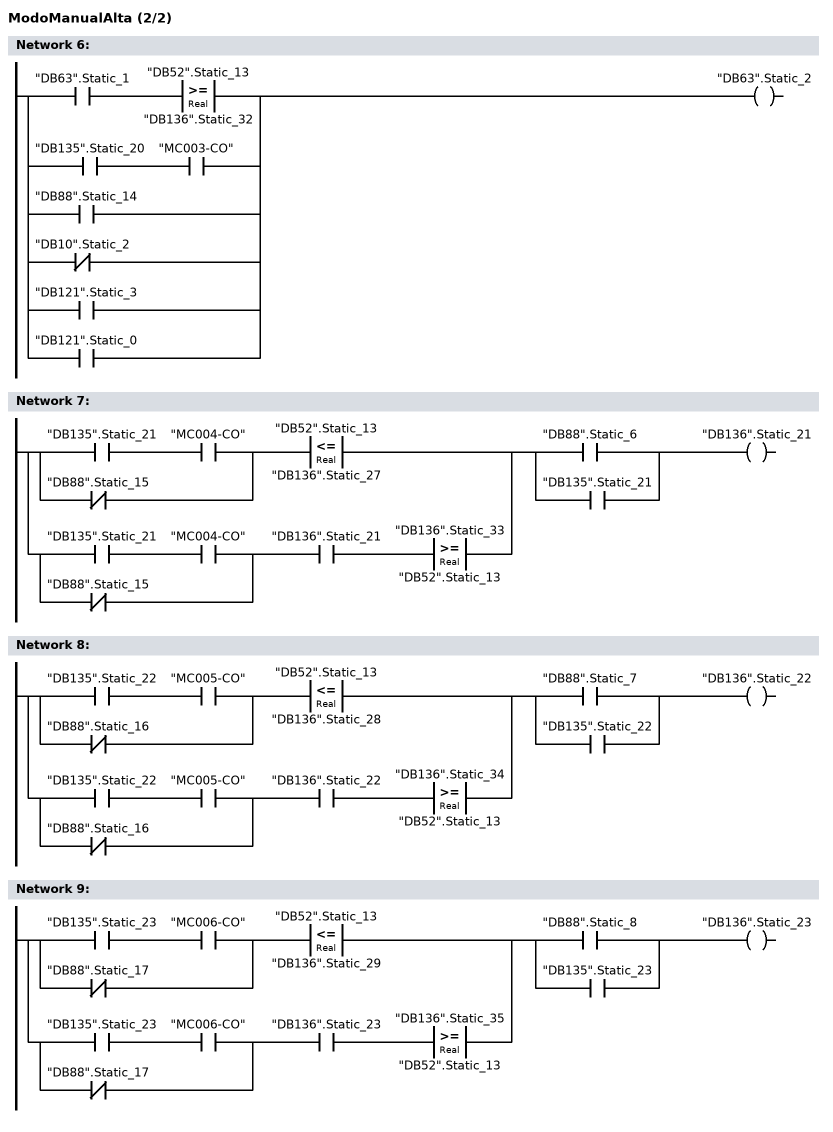
   "DB63".Static_2 := ("DB63".Static_1 AND ("DB52".Static_13 >= "DB136".Static_32)) OR "DB88".Static_14 OR ("DB135".Static_20 AND "MC003-CO") OR NOT "DB10".Static_2 OR "DB121".Static_3 OR "DB121".Static_0;
END_REGION

REGION Network 7
   "DB136".Static_21 := (((NOT "DB88".Static_15 OR ("DB135".Static_21 AND "MC004-CO")) AND ("DB52".Static_13 <= "DB136".Static_27)) OR ((NOT "DB88".Static_15 OR ("DB135".Static_21 AND "MC004-CO")) AND "DB136".Static_21 AND ("DB136".Static_33 >= "DB52".Static_13))) AND ("DB88".Static_6 OR "DB135".Static_21);
END_REGION

REGION Network 8
   "DB136".Static_22 := (((NOT "DB88".Static_16 OR ("DB135".Static_22 AND "MC005-CO")) AND ("DB52".Static_13 <= "DB136".Static_28)) OR ((NOT "DB88".Static_16 OR ("DB135".Static_22 AND "MC005-CO")) AND "DB136".Static_22 AND ("DB136".Static_34 >= "DB52".Static_13))) AND ("DB88".Static_7 OR "DB135".Static_22);
END_REGION

REGION Network 9
   "DB136".Static_23 := (((NOT "DB88".Static_17 OR ("DB135".Static_23 AND "MC006-CO")) AND ("DB52".Static_13 <= "DB136".Static_29)) OR ((NOT "DB88".Static_17 OR ("DB135".Static_23 AND "MC006-CO")) AND "DB136".Static_23 AND ("DB136".Static_35 >= "DB52".Static_13))) AND ("DB88".Static_8 OR "DB135".Static_23);
END_REGION
END_FUNCTION

// folder: Compresores/Alta/Maquina de Estados

FUNCTION "LogMaqEstGeneral" : Void   // FC35, LAD
{ S7_Optimized_Access := 'FALSE' }
VERSION : 0.1
BEGIN

REGION Network 1
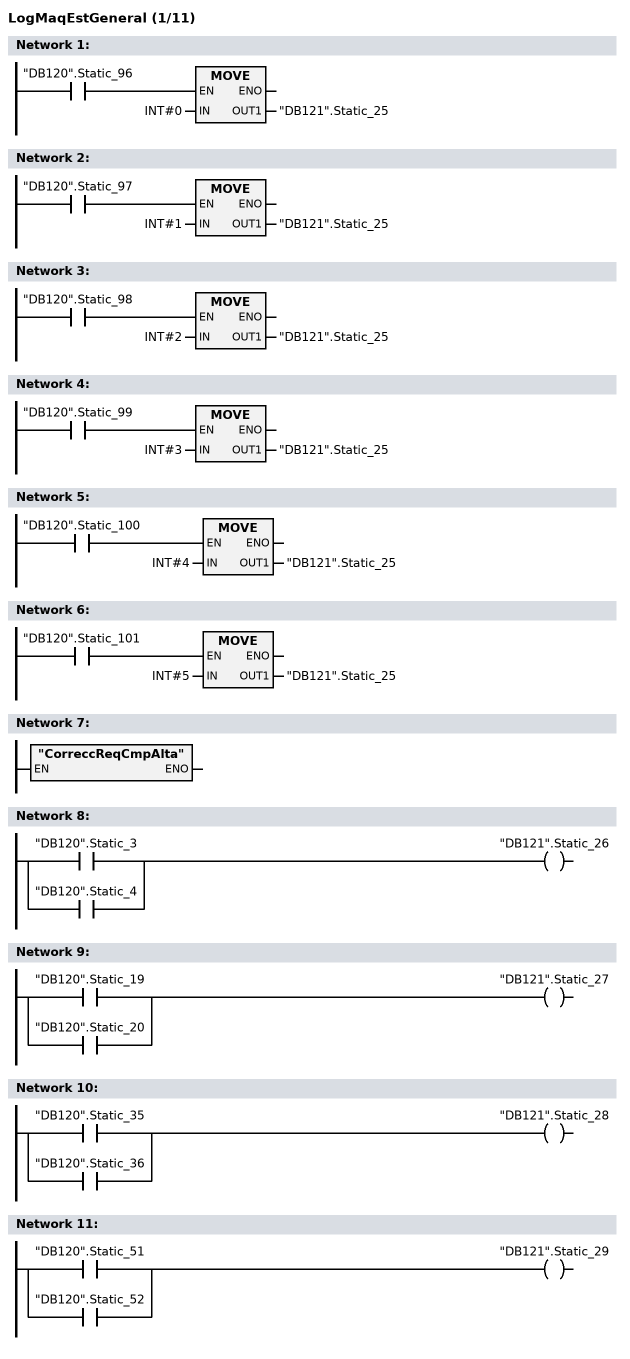
   RUNG wire#powerrail
      Contact( "DB120".Static_96 )
      { S7_GenerateENO := "TRUE" } Move(in := INT#0, out1 => "DB121".Static_25)
   END_RUNG
   // the same network as SCL:
   IF "DB120".Static_96 THEN "DB121".Static_25 := INT#0; END_IF;
END_REGION

REGION Network 2
   RUNG wire#powerrail
      Contact( "DB120".Static_97 )
      { S7_GenerateENO := "TRUE" } Move(in := INT#1, out1 => "DB121".Static_25)
   END_RUNG
   // the same network as SCL:
   IF "DB120".Static_97 THEN "DB121".Static_25 := INT#1; END_IF;
END_REGION

REGION Network 3
   RUNG wire#powerrail
      Contact( "DB120".Static_98 )
      { S7_GenerateENO := "TRUE" } Move(in := INT#2, out1 => "DB121".Static_25)
   END_RUNG
   // the same network as SCL:
   IF "DB120".Static_98 THEN "DB121".Static_25 := INT#2; END_IF;
END_REGION

REGION Network 4
   RUNG wire#powerrail
      Contact( "DB120".Static_99 )
      { S7_GenerateENO := "TRUE" } Move(in := INT#3, out1 => "DB121".Static_25)
   END_RUNG
   // the same network as SCL:
   IF "DB120".Static_99 THEN "DB121".Static_25 := INT#3; END_IF;
END_REGION

REGION Network 5
   RUNG wire#powerrail
      Contact( "DB120".Static_100 )
      { S7_GenerateENO := "TRUE" } Move(in := INT#4, out1 => "DB121".Static_25)
   END_RUNG
   // the same network as SCL:
   IF "DB120".Static_100 THEN "DB121".Static_25 := INT#4; END_IF;
END_REGION

REGION Network 6
   RUNG wire#powerrail
      Contact( "DB120".Static_101 )
      { S7_GenerateENO := "TRUE" } Move(in := INT#5, out1 => "DB121".Static_25)
   END_RUNG
   // the same network as SCL:
   IF "DB120".Static_101 THEN "DB121".Static_25 := INT#5; END_IF;
END_REGION

REGION Network 7
   RUNG wire#powerrail
      "CorreccReqCmpAlta"()
   END_RUNG
   // the same network as SCL:
   "CorreccReqCmpAlta"();
END_REGION

REGION Network 8
   RUNG wire#powerrail
      Contact( "DB120".Static_3 )
      wire#w1
      Coil( "DB121".Static_26 )
   END_RUNG
   RUNG wire#powerrail
      Contact( "DB120".Static_4 )
   END_RUNG wire#w1
   // the same network as SCL:
   "DB121".Static_26 := "DB120".Static_3 OR "DB120".Static_4;
END_REGION

REGION Network 9
   RUNG wire#powerrail
      Contact( "DB120".Static_19 )
      wire#w1
      Coil( "DB121".Static_27 )
   END_RUNG
   RUNG wire#powerrail
      Contact( "DB120".Static_20 )
   END_RUNG wire#w1
   // the same network as SCL:
   "DB121".Static_27 := "DB120".Static_19 OR "DB120".Static_20;
END_REGION

REGION Network 10
   RUNG wire#powerrail
      Contact( "DB120".Static_35 )
      wire#w1
      Coil( "DB121".Static_28 )
   END_RUNG
   RUNG wire#powerrail
      Contact( "DB120".Static_36 )
   END_RUNG wire#w1
   // the same network as SCL:
   "DB121".Static_28 := "DB120".Static_35 OR "DB120".Static_36;
END_REGION

REGION Network 11
   RUNG wire#powerrail
      Contact( "DB120".Static_51 )
      wire#w1
      Coil( "DB121".Static_29 )
   END_RUNG
   RUNG wire#powerrail
      Contact( "DB120".Static_52 )
   END_RUNG wire#w1
   // the same network as SCL:
   "DB121".Static_29 := "DB120".Static_51 OR "DB120".Static_52;
END_REGION

REGION Network 12
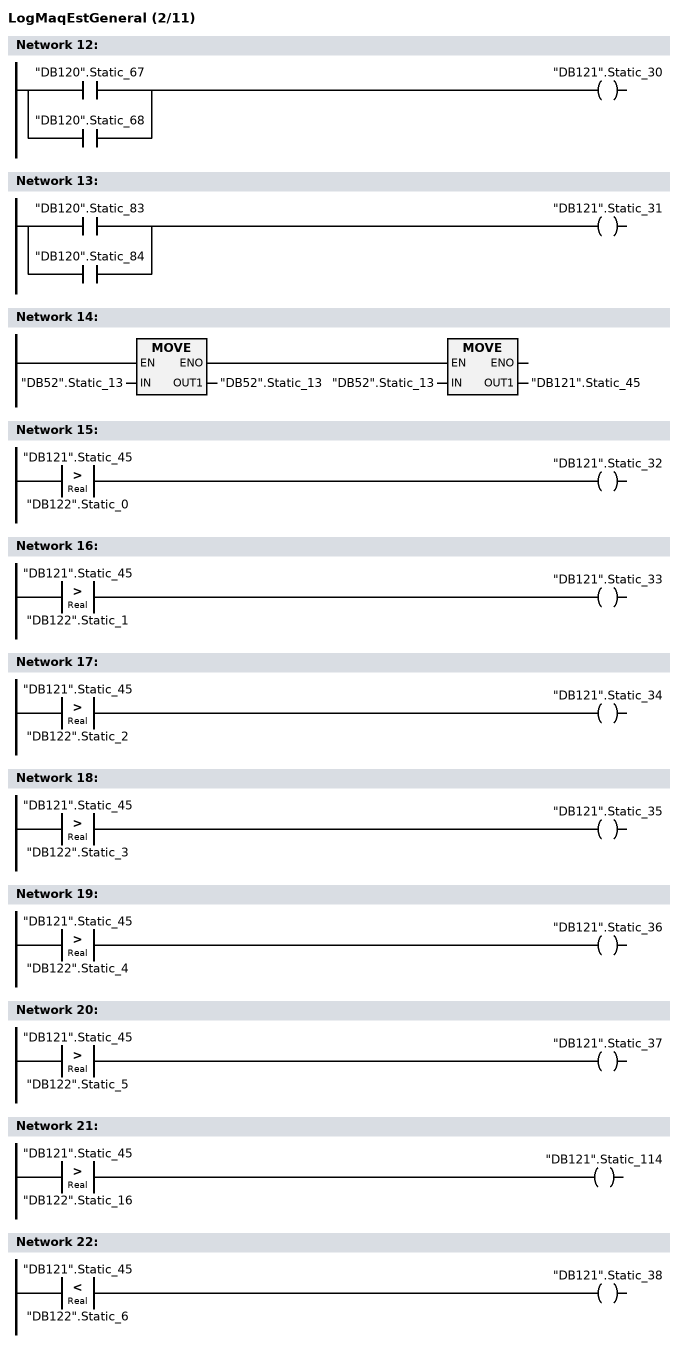
   RUNG wire#powerrail
      Contact( "DB120".Static_67 )
      wire#w1
      Coil( "DB121".Static_30 )
   END_RUNG
   RUNG wire#powerrail
      Contact( "DB120".Static_68 )
   END_RUNG wire#w1
   // the same network as SCL:
   "DB121".Static_30 := "DB120".Static_67 OR "DB120".Static_68;
END_REGION

REGION Network 13
   RUNG wire#powerrail
      Contact( "DB120".Static_83 )
      wire#w1
      Coil( "DB121".Static_31 )
   END_RUNG
   RUNG wire#powerrail
      Contact( "DB120".Static_84 )
   END_RUNG wire#w1
   // the same network as SCL:
   "DB121".Static_31 := "DB120".Static_83 OR "DB120".Static_84;
END_REGION

REGION Network 14
   RUNG wire#powerrail
      { S7_GenerateENO := "TRUE" } Move(in := "DB52".Static_13, out1 => "DB52".Static_13)
      { S7_GenerateENO := "TRUE" } Move(in := "DB52".Static_13, out1 => "DB121".Static_45)
   END_RUNG
   // the same network as SCL:
   // ENO of a box is taken as its EN; it also drops when the box reports an error
   "DB52".Static_13 := "DB52".Static_13;
   "DB121".Static_45 := "DB52".Static_13;
END_REGION

REGION Network 15
   RUNG wire#powerrail
      { S7_Templates := "SrcType := Real" } GT_Contact(in1 := "DB121".Static_45, in2 := "DB122".Static_0)
      Coil( "DB121".Static_32 )
   END_RUNG
   // the same network as SCL:
   "DB121".Static_32 := "DB121".Static_45 > "DB122".Static_0;
END_REGION

REGION Network 16
   RUNG wire#powerrail
      { S7_Templates := "SrcType := Real" } GT_Contact(in1 := "DB121".Static_45, in2 := "DB122".Static_1)
      Coil( "DB121".Static_33 )
   END_RUNG
   // the same network as SCL:
   "DB121".Static_33 := "DB121".Static_45 > "DB122".Static_1;
END_REGION

REGION Network 17
   RUNG wire#powerrail
      { S7_Templates := "SrcType := Real" } GT_Contact(in1 := "DB121".Static_45, in2 := "DB122".Static_2)
      Coil( "DB121".Static_34 )
   END_RUNG
   // the same network as SCL:
   "DB121".Static_34 := "DB121".Static_45 > "DB122".Static_2;
END_REGION

REGION Network 18
   RUNG wire#powerrail
      { S7_Templates := "SrcType := Real" } GT_Contact(in1 := "DB121".Static_45, in2 := "DB122".Static_3)
      Coil( "DB121".Static_35 )
   END_RUNG
   // the same network as SCL:
   "DB121".Static_35 := "DB121".Static_45 > "DB122".Static_3;
END_REGION

REGION Network 19
   RUNG wire#powerrail
      { S7_Templates := "SrcType := Real" } GT_Contact(in1 := "DB121".Static_45, in2 := "DB122".Static_4)
      Coil( "DB121".Static_36 )
   END_RUNG
   // the same network as SCL:
   "DB121".Static_36 := "DB121".Static_45 > "DB122".Static_4;
END_REGION

REGION Network 20
   RUNG wire#powerrail
      { S7_Templates := "SrcType := Real" } GT_Contact(in1 := "DB121".Static_45, in2 := "DB122".Static_5)
      Coil( "DB121".Static_37 )
   END_RUNG
   // the same network as SCL:
   "DB121".Static_37 := "DB121".Static_45 > "DB122".Static_5;
END_REGION

REGION Network 21
   RUNG wire#powerrail
      { S7_Templates := "SrcType := Real" } GT_Contact(in1 := "DB121".Static_45, in2 := "DB122".Static_16)
      Coil( "DB121".Static_114 )
   END_RUNG
   // the same network as SCL:
   "DB121".Static_114 := "DB121".Static_45 > "DB122".Static_16;
END_REGION

REGION Network 22
   RUNG wire#powerrail
      { S7_Templates := "SrcType := Real" } LT_Contact(in1 := "DB121".Static_45, in2 := "DB122".Static_6)
      Coil( "DB121".Static_38 )
   END_RUNG
   // the same network as SCL:
   "DB121".Static_38 := "DB121".Static_45 < "DB122".Static_6;
END_REGION

REGION Network 23
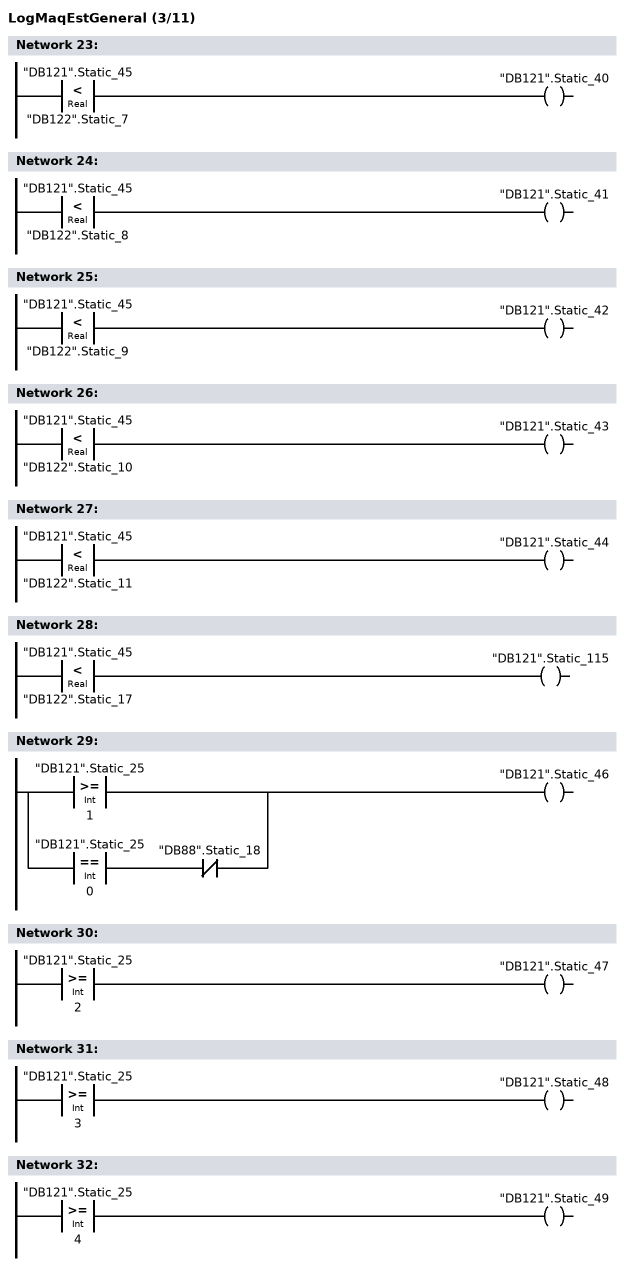
   RUNG wire#powerrail
      { S7_Templates := "SrcType := Real" } LT_Contact(in1 := "DB121".Static_45, in2 := "DB122".Static_7)
      Coil( "DB121".Static_40 )
   END_RUNG
   // the same network as SCL:
   "DB121".Static_40 := "DB121".Static_45 < "DB122".Static_7;
END_REGION

REGION Network 24
   RUNG wire#powerrail
      { S7_Templates := "SrcType := Real" } LT_Contact(in1 := "DB121".Static_45, in2 := "DB122".Static_8)
      Coil( "DB121".Static_41 )
   END_RUNG
   // the same network as SCL:
   "DB121".Static_41 := "DB121".Static_45 < "DB122".Static_8;
END_REGION

REGION Network 25
   RUNG wire#powerrail
      { S7_Templates := "SrcType := Real" } LT_Contact(in1 := "DB121".Static_45, in2 := "DB122".Static_9)
      Coil( "DB121".Static_42 )
   END_RUNG
   // the same network as SCL:
   "DB121".Static_42 := "DB121".Static_45 < "DB122".Static_9;
END_REGION

REGION Network 26
   RUNG wire#powerrail
      { S7_Templates := "SrcType := Real" } LT_Contact(in1 := "DB121".Static_45, in2 := "DB122".Static_10)
      Coil( "DB121".Static_43 )
   END_RUNG
   // the same network as SCL:
   "DB121".Static_43 := "DB121".Static_45 < "DB122".Static_10;
END_REGION

REGION Network 27
   RUNG wire#powerrail
      { S7_Templates := "SrcType := Real" } LT_Contact(in1 := "DB121".Static_45, in2 := "DB122".Static_11)
      Coil( "DB121".Static_44 )
   END_RUNG
   // the same network as SCL:
   "DB121".Static_44 := "DB121".Static_45 < "DB122".Static_11;
END_REGION

REGION Network 28
   RUNG wire#powerrail
      { S7_Templates := "SrcType := Real" } LT_Contact(in1 := "DB121".Static_45, in2 := "DB122".Static_17)
      Coil( "DB121".Static_115 )
   END_RUNG
   // the same network as SCL:
   "DB121".Static_115 := "DB121".Static_45 < "DB122".Static_17;
END_REGION

REGION Network 29
   RUNG wire#powerrail
      { S7_Templates := "SrcType := Int" } GE_Contact(in1 := "DB121".Static_25, in2 := 1)
      wire#w1
      Coil( "DB121".Static_46 )
   END_RUNG
   RUNG wire#powerrail
      { S7_Templates := "SrcType := Int" } EQ_Contact(in1 := "DB121".Static_25, in2 := 0)
      I_Contact( "DB88".Static_18 )
   END_RUNG wire#w1
   // the same network as SCL:
   "DB121".Static_46 := ("DB121".Static_25 >= 1) OR (("DB121".Static_25 = 0) AND NOT "DB88".Static_18);
END_REGION

REGION Network 30
   RUNG wire#powerrail
      { S7_Templates := "SrcType := Int" } GE_Contact(in1 := "DB121".Static_25, in2 := 2)
      Coil( "DB121".Static_47 )
   END_RUNG
   // the same network as SCL:
   "DB121".Static_47 := "DB121".Static_25 >= 2;
END_REGION

REGION Network 31
   RUNG wire#powerrail
      { S7_Templates := "SrcType := Int" } GE_Contact(in1 := "DB121".Static_25, in2 := 3)
      Coil( "DB121".Static_48 )
   END_RUNG
   // the same network as SCL:
   "DB121".Static_48 := "DB121".Static_25 >= 3;
END_REGION

REGION Network 32
   RUNG wire#powerrail
      { S7_Templates := "SrcType := Int" } GE_Contact(in1 := "DB121".Static_25, in2 := 4)
      Coil( "DB121".Static_49 )
   END_RUNG
   // the same network as SCL:
   "DB121".Static_49 := "DB121".Static_25 >= 4;
END_REGION

REGION Network 33
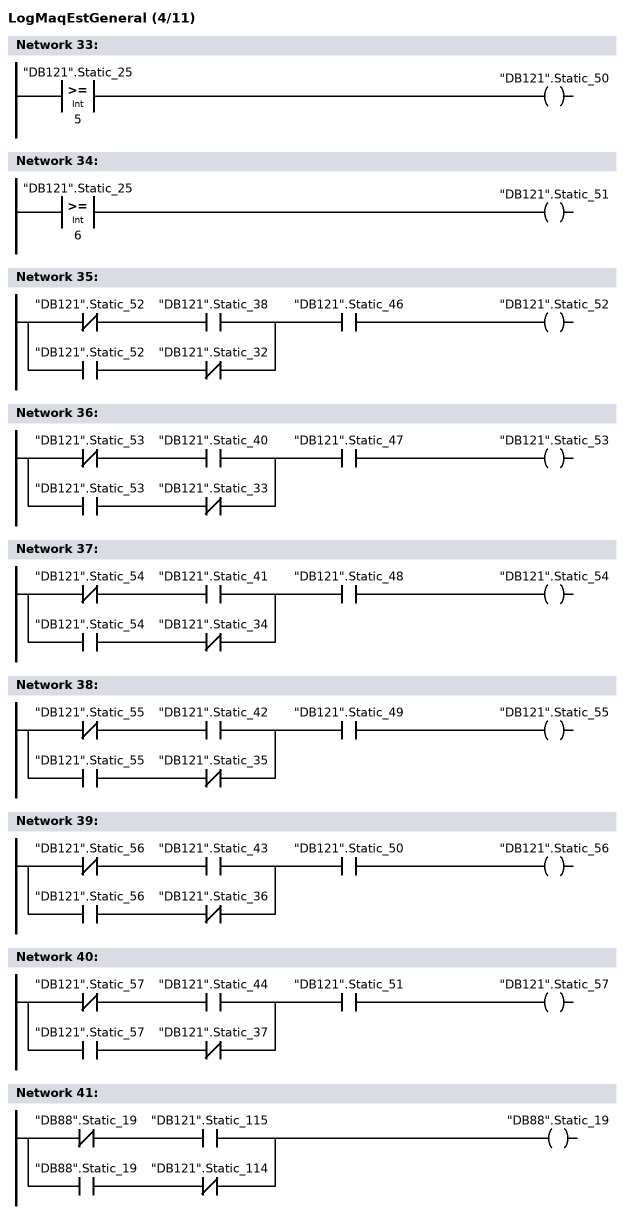
   RUNG wire#powerrail
      { S7_Templates := "SrcType := Int" } GE_Contact(in1 := "DB121".Static_25, in2 := 5)
      Coil( "DB121".Static_50 )
   END_RUNG
   // the same network as SCL:
   "DB121".Static_50 := "DB121".Static_25 >= 5;
END_REGION

REGION Network 34
   RUNG wire#powerrail
      { S7_Templates := "SrcType := Int" } GE_Contact(in1 := "DB121".Static_25, in2 := 6)
      Coil( "DB121".Static_51 )
   END_RUNG
   // the same network as SCL:
   "DB121".Static_51 := "DB121".Static_25 >= 6;
END_REGION

REGION Network 35
   RUNG wire#powerrail
      I_Contact( "DB121".Static_52 )
      Contact( "DB121".Static_38 )
      wire#w1
      Contact( "DB121".Static_46 )
      Coil( "DB121".Static_52 )
   END_RUNG
   RUNG wire#powerrail
      Contact( "DB121".Static_52 )
      I_Contact( "DB121".Static_32 )
   END_RUNG wire#w1
   // the same network as SCL:
   "DB121".Static_52 := ((NOT "DB121".Static_52 AND "DB121".Static_38) OR ("DB121".Static_52 AND NOT "DB121".Static_32)) AND "DB121".Static_46;
END_REGION

REGION Network 36
   RUNG wire#powerrail
      I_Contact( "DB121".Static_53 )
      Contact( "DB121".Static_40 )
      wire#w1
      Contact( "DB121".Static_47 )
      Coil( "DB121".Static_53 )
   END_RUNG
   RUNG wire#powerrail
      Contact( "DB121".Static_53 )
      I_Contact( "DB121".Static_33 )
   END_RUNG wire#w1
   // the same network as SCL:
   "DB121".Static_53 := ((NOT "DB121".Static_53 AND "DB121".Static_40) OR ("DB121".Static_53 AND NOT "DB121".Static_33)) AND "DB121".Static_47;
END_REGION

REGION Network 37
   RUNG wire#powerrail
      I_Contact( "DB121".Static_54 )
      Contact( "DB121".Static_41 )
      wire#w1
      Contact( "DB121".Static_48 )
      Coil( "DB121".Static_54 )
   END_RUNG
   RUNG wire#powerrail
      Contact( "DB121".Static_54 )
      I_Contact( "DB121".Static_34 )
   END_RUNG wire#w1
   // the same network as SCL:
   "DB121".Static_54 := ((NOT "DB121".Static_54 AND "DB121".Static_41) OR ("DB121".Static_54 AND NOT "DB121".Static_34)) AND "DB121".Static_48;
END_REGION

REGION Network 38
   RUNG wire#powerrail
      I_Contact( "DB121".Static_55 )
      Contact( "DB121".Static_42 )
      wire#w1
      Contact( "DB121".Static_49 )
      Coil( "DB121".Static_55 )
   END_RUNG
   RUNG wire#powerrail
      Contact( "DB121".Static_55 )
      I_Contact( "DB121".Static_35 )
   END_RUNG wire#w1
   // the same network as SCL:
   "DB121".Static_55 := ((NOT "DB121".Static_55 AND "DB121".Static_42) OR ("DB121".Static_55 AND NOT "DB121".Static_35)) AND "DB121".Static_49;
END_REGION

REGION Network 39
   RUNG wire#powerrail
      I_Contact( "DB121".Static_56 )
      Contact( "DB121".Static_43 )
      wire#w1
      Contact( "DB121".Static_50 )
      Coil( "DB121".Static_56 )
   END_RUNG
   RUNG wire#powerrail
      Contact( "DB121".Static_56 )
      I_Contact( "DB121".Static_36 )
   END_RUNG wire#w1
   // the same network as SCL:
   "DB121".Static_56 := ((NOT "DB121".Static_56 AND "DB121".Static_43) OR ("DB121".Static_56 AND NOT "DB121".Static_36)) AND "DB121".Static_50;
END_REGION

REGION Network 40
   RUNG wire#powerrail
      I_Contact( "DB121".Static_57 )
      Contact( "DB121".Static_44 )
      wire#w1
      Contact( "DB121".Static_51 )
      Coil( "DB121".Static_57 )
   END_RUNG
   RUNG wire#powerrail
      Contact( "DB121".Static_57 )
      I_Contact( "DB121".Static_37 )
   END_RUNG wire#w1
   // the same network as SCL:
   "DB121".Static_57 := ((NOT "DB121".Static_57 AND "DB121".Static_44) OR ("DB121".Static_57 AND NOT "DB121".Static_37)) AND "DB121".Static_51;
END_REGION

REGION Network 41
   RUNG wire#powerrail
      I_Contact( "DB88".Static_19 )
      Contact( "DB121".Static_115 )
      wire#w1
      Coil( "DB88".Static_19 )
   END_RUNG
   RUNG wire#powerrail
      Contact( "DB88".Static_19 )
      I_Contact( "DB121".Static_114 )
   END_RUNG wire#w1
   // the same network as SCL:
   "DB88".Static_19 := (NOT "DB88".Static_19 AND "DB121".Static_115) OR ("DB88".Static_19 AND NOT "DB121".Static_114);
END_REGION

REGION Network 42
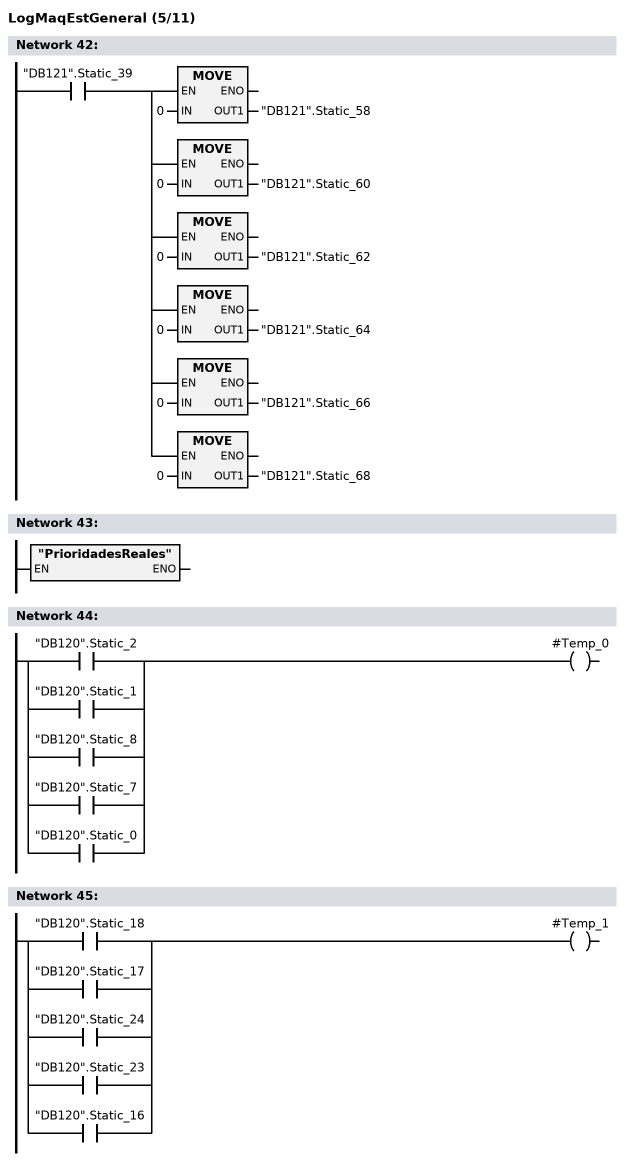
   RUNG wire#powerrail
      Contact( "DB121".Static_39 )
      wire#w1
      { S7_GenerateENO := "TRUE" } Move(in := 0, out1 => "DB121".Static_58)
   END_RUNG
   RUNG wire#w1
      { S7_GenerateENO := "TRUE" } Move(in := 0, out1 => "DB121".Static_60)
   END_RUNG
   RUNG wire#w1
      { S7_GenerateENO := "TRUE" } Move(in := 0, out1 => "DB121".Static_62)
   END_RUNG
   RUNG wire#w1
      { S7_GenerateENO := "TRUE" } Move(in := 0, out1 => "DB121".Static_64)
   END_RUNG
   RUNG wire#w1
      { S7_GenerateENO := "TRUE" } Move(in := 0, out1 => "DB121".Static_66)
   END_RUNG
   RUNG wire#w1
      { S7_GenerateENO := "TRUE" } Move(in := 0, out1 => "DB121".Static_68)
   END_RUNG
   // the same network as SCL:
   IF "DB121".Static_39 THEN
       "DB121".Static_58 := 0;
       "DB121".Static_60 := 0;
       "DB121".Static_62 := 0;
       "DB121".Static_64 := 0;
       "DB121".Static_66 := 0;
       "DB121".Static_68 := 0;
   END_IF;
END_REGION

REGION Network 43
   RUNG wire#powerrail
      "PrioridadesReales"()
   END_RUNG
   // the same network as SCL:
   "PrioridadesReales"();
END_REGION

REGION Network 44
   RUNG wire#powerrail
      Contact( "DB120".Static_2 )
      wire#w1
      Coil( #Temp_0 )
   END_RUNG
   RUNG wire#powerrail
      Contact( "DB120".Static_1 )
   END_RUNG wire#w1
   RUNG wire#powerrail
      Contact( "DB120".Static_8 )
   END_RUNG wire#w1
   RUNG wire#powerrail
      Contact( "DB120".Static_7 )
   END_RUNG wire#w1
   RUNG wire#powerrail
      Contact( "DB120".Static_0 )
   END_RUNG wire#w1
   // the same network as SCL:
   #Temp_0 := "DB120".Static_2 OR "DB120".Static_1 OR "DB120".Static_8 OR "DB120".Static_7 OR "DB120".Static_0;
END_REGION

REGION Network 45
   RUNG wire#powerrail
      Contact( "DB120".Static_18 )
      wire#w1
      Coil( #Temp_1 )
   END_RUNG
   RUNG wire#powerrail
      Contact( "DB120".Static_17 )
   END_RUNG wire#w1
   RUNG wire#powerrail
      Contact( "DB120".Static_24 )
   END_RUNG wire#w1
   RUNG wire#powerrail
      Contact( "DB120".Static_23 )
   END_RUNG wire#w1
   RUNG wire#powerrail
      Contact( "DB120".Static_16 )
   END_RUNG wire#w1
   // the same network as SCL:
   #Temp_1 := "DB120".Static_18 OR "DB120".Static_17 OR "DB120".Static_24 OR "DB120".Static_23 OR "DB120".Static_16;
END_REGION

REGION Network 46
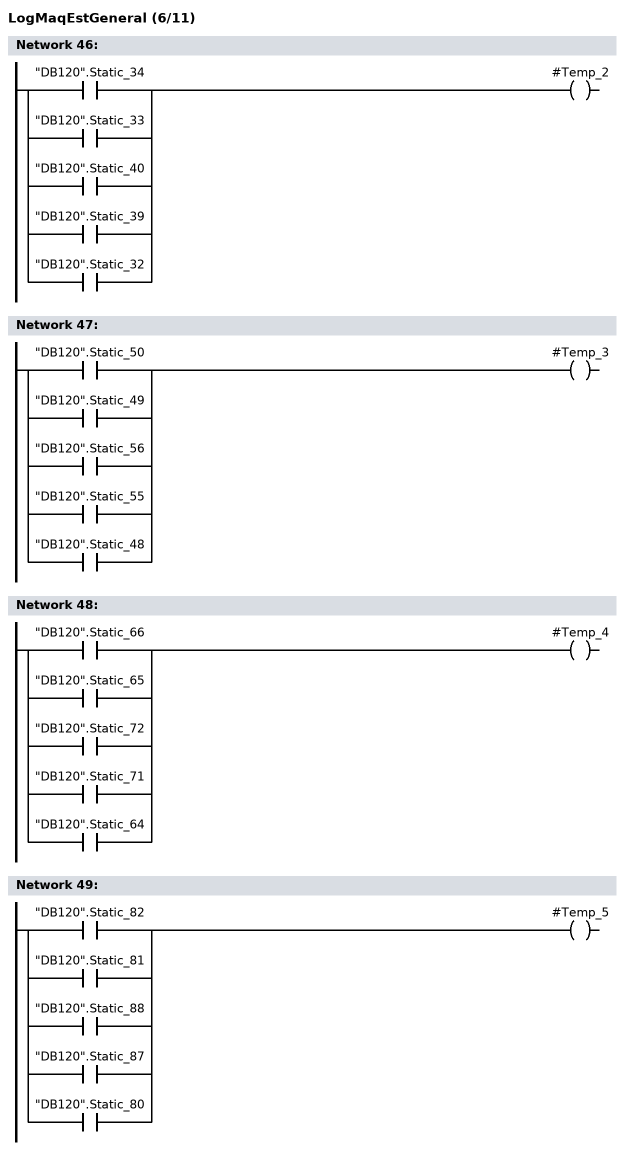
   RUNG wire#powerrail
      Contact( "DB120".Static_34 )
      wire#w1
      Coil( #Temp_2 )
   END_RUNG
   RUNG wire#powerrail
      Contact( "DB120".Static_33 )
   END_RUNG wire#w1
   RUNG wire#powerrail
      Contact( "DB120".Static_40 )
   END_RUNG wire#w1
   RUNG wire#powerrail
      Contact( "DB120".Static_39 )
   END_RUNG wire#w1
   RUNG wire#powerrail
      Contact( "DB120".Static_32 )
   END_RUNG wire#w1
   // the same network as SCL:
   #Temp_2 := "DB120".Static_34 OR "DB120".Static_33 OR "DB120".Static_40 OR "DB120".Static_39 OR "DB120".Static_32;
END_REGION

REGION Network 47
   RUNG wire#powerrail
      Contact( "DB120".Static_50 )
      wire#w1
      Coil( #Temp_3 )
   END_RUNG
   RUNG wire#powerrail
      Contact( "DB120".Static_49 )
   END_RUNG wire#w1
   RUNG wire#powerrail
      Contact( "DB120".Static_56 )
   END_RUNG wire#w1
   RUNG wire#powerrail
      Contact( "DB120".Static_55 )
   END_RUNG wire#w1
   RUNG wire#powerrail
      Contact( "DB120".Static_48 )
   END_RUNG wire#w1
   // the same network as SCL:
   #Temp_3 := "DB120".Static_50 OR "DB120".Static_49 OR "DB120".Static_56 OR "DB120".Static_55 OR "DB120".Static_48;
END_REGION

REGION Network 48
   RUNG wire#powerrail
      Contact( "DB120".Static_66 )
      wire#w1
      Coil( #Temp_4 )
   END_RUNG
   RUNG wire#powerrail
      Contact( "DB120".Static_65 )
   END_RUNG wire#w1
   RUNG wire#powerrail
      Contact( "DB120".Static_72 )
   END_RUNG wire#w1
   RUNG wire#powerrail
      Contact( "DB120".Static_71 )
   END_RUNG wire#w1
   RUNG wire#powerrail
      Contact( "DB120".Static_64 )
   END_RUNG wire#w1
   // the same network as SCL:
   #Temp_4 := "DB120".Static_66 OR "DB120".Static_65 OR "DB120".Static_72 OR "DB120".Static_71 OR "DB120".Static_64;
END_REGION

REGION Network 49
   RUNG wire#powerrail
      Contact( "DB120".Static_82 )
      wire#w1
      Coil( #Temp_5 )
   END_RUNG
   RUNG wire#powerrail
      Contact( "DB120".Static_81 )
   END_RUNG wire#w1
   RUNG wire#powerrail
      Contact( "DB120".Static_88 )
   END_RUNG wire#w1
   RUNG wire#powerrail
      Contact( "DB120".Static_87 )
   END_RUNG wire#w1
   RUNG wire#powerrail
      Contact( "DB120".Static_80 )
   END_RUNG wire#w1
   // the same network as SCL:
   #Temp_5 := "DB120".Static_82 OR "DB120".Static_81 OR "DB120".Static_88 OR "DB120".Static_87 OR "DB120".Static_80;
END_REGION

REGION Network 50 (STL)
         A     #Temp_0;
         A(;
         A     "DB121".Static_46;
         A(;
         L     "DB121".Static_58;
         L     1;
         ==R;
         );
         O;
         A     "DB121".Static_47;
         A(;
         L     "DB121".Static_58;
         L     2;
         ==R;
         );
         O;
         A     "DB121".Static_48;
         A(;
         L     "DB121".Static_58;
         L     3;
         ==R;
         );
         O;
         A     "DB121".Static_49;
         A(;
         L     "DB121".Static_58;
         L     4;
         ==R;
         );
         O;
         A     "DB121".Static_50;
         A(;
         L     "DB121".Static_58;
         L     5;
         ==R;
         );
         O;
         A     "DB121".Static_51;
         A(;
         L     "DB121".Static_58;
         L     6;
         ==R;
         );
         );
         =     "DB121".Static_70;
END_REGION

REGION Network 51 (STL)
         A     #Temp_1;
         A(;
         A     "DB121".Static_46;
         A(;
         L     "DB121".Static_60;
         L     1;
         ==R;
         );
         O;
         A     "DB121".Static_47;
         A(;
         L     "DB121".Static_60;
         L     2;
         ==R;
         );
         O;
         A     "DB121".Static_48;
         A(;
         L     "DB121".Static_60;
         L     3;
         ==R;
         );
         O;
         A     "DB121".Static_49;
         A(;
         L     "DB121".Static_60;
         L     4;
         ==R;
         );
         O;
         A     "DB121".Static_50;
         A(;
         L     "DB121".Static_60;
         L     5;
         ==R;
         );
         O;
         A     "DB121".Static_51;
         A(;
         L     "DB121".Static_60;
         L     6;
         ==R;
         );
         );
         =     "DB121".Static_71;
END_REGION

REGION Network 52 (STL)
         A     #Temp_2;
         A(;
         A     "DB121".Static_46;
         A(;
         L     "DB121".Static_62;
         L     1;
         ==R;
         );
         O;
         A     "DB121".Static_47;
         A(;
         L     "DB121".Static_62;
         L     2;
         ==R;
         );
         O;
         A     "DB121".Static_48;
         A(;
         L     "DB121".Static_62;
         L     3;
         ==R;
         );
         O;
         A     "DB121".Static_49;
         A(;
         L     "DB121".Static_62;
         L     4;
         ==R;
         );
         O;
         A     "DB121".Static_50;
         A(;
         L     "DB121".Static_62;
         L     5;
         ==R;
         );
         O;
         A     "DB121".Static_51;
         A(;
         L     "DB121".Static_62;
         L     6;
         ==R;
         );
         );
         =     "DB121".Static_72;
END_REGION

REGION Network 53 (STL)
         A     #Temp_3;
         A(;
         A     "DB121".Static_46;
         A(;
         L     "DB121".Static_64;
         L     1;
         ==R;
         );
         O;
         A     "DB121".Static_47;
         A(;
         L     "DB121".Static_64;
         L     2;
         ==R;
         );
         O;
         A     "DB121".Static_48;
         A(;
         L     "DB121".Static_64;
         L     3;
         ==R;
         );
         O;
         A     "DB121".Static_49;
         A(;
         L     "DB121".Static_64;
         L     4;
         ==R;
         );
         O;
         A     "DB121".Static_50;
         A(;
         L     "DB121".Static_64;
         L     5;
         ==R;
         );
         O;
         A     "DB121".Static_51;
         A(;
         L     "DB121".Static_64;
         L     6;
         ==R;
         );
         );
         =     "DB121".Static_73;
END_REGION

REGION Network 54 (STL)
         A     #Temp_4;
         A(;
         A     "DB121".Static_46;
         A(;
         L     "DB121".Static_66;
         L     1;
         ==R;
         );
         O;
         A     "DB121".Static_47;
         A(;
         L     "DB121".Static_66;
         L     2;
         ==R;
         );
         O;
         A     "DB121".Static_48;
         A(;
         L     "DB121".Static_66;
         L     3;
         ==R;
         );
         O;
         A     "DB121".Static_49;
         A(;
         L     "DB121".Static_66;
         L     4;
         ==R;
         );
         O;
         A     "DB121".Static_50;
         A(;
         L     "DB121".Static_66;
         L     5;
         ==R;
         );
         O;
         A     "DB121".Static_51;
         A(;
         L     "DB121".Static_66;
         L     6;
         ==R;
         );
         );
         =     "DB121".Static_74;
END_REGION

REGION Network 55 (STL)
         A     #Temp_5;
         A(;
         A     "DB121".Static_46;
         A(;
         L     "DB121".Static_68;
         L     1;
         ==R;
         );
         O;
         A     "DB121".Static_47;
         A(;
         L     "DB121".Static_68;
         L     2;
         ==R;
         );
         O;
         A     "DB121".Static_48;
         A(;
         L     "DB121".Static_68;
         L     3;
         ==R;
         );
         O;
         A     "DB121".Static_49;
         A(;
         L     "DB121".Static_68;
         L     4;
         ==R;
         );
         O;
         A     "DB121".Static_50;
         A(;
         L     "DB121".Static_68;
         L     5;
         ==R;
         );
         O;
         A     "DB121".Static_51;
         A(;
         L     "DB121".Static_68;
         L     6;
         ==R;
         );
         );
         =     "DB121".Static_75;
END_REGION

REGION Network 56
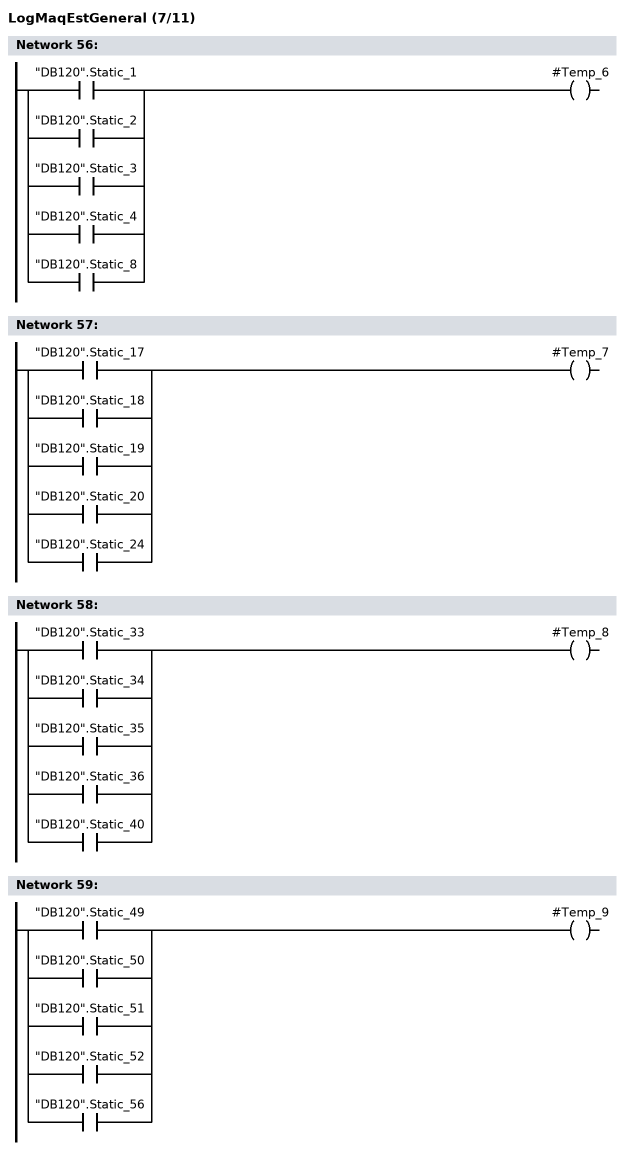
   RUNG wire#powerrail
      Contact( "DB120".Static_1 )
      wire#w1
      Coil( #Temp_6 )
   END_RUNG
   RUNG wire#powerrail
      Contact( "DB120".Static_2 )
   END_RUNG wire#w1
   RUNG wire#powerrail
      Contact( "DB120".Static_3 )
   END_RUNG wire#w1
   RUNG wire#powerrail
      Contact( "DB120".Static_4 )
   END_RUNG wire#w1
   RUNG wire#powerrail
      Contact( "DB120".Static_8 )
   END_RUNG wire#w1
   // the same network as SCL:
   #Temp_6 := "DB120".Static_1 OR "DB120".Static_2 OR "DB120".Static_3 OR "DB120".Static_4 OR "DB120".Static_8;
END_REGION

REGION Network 57
   RUNG wire#powerrail
      Contact( "DB120".Static_17 )
      wire#w1
      Coil( #Temp_7 )
   END_RUNG
   RUNG wire#powerrail
      Contact( "DB120".Static_18 )
   END_RUNG wire#w1
   RUNG wire#powerrail
      Contact( "DB120".Static_19 )
   END_RUNG wire#w1
   RUNG wire#powerrail
      Contact( "DB120".Static_20 )
   END_RUNG wire#w1
   RUNG wire#powerrail
      Contact( "DB120".Static_24 )
   END_RUNG wire#w1
   // the same network as SCL:
   #Temp_7 := "DB120".Static_17 OR "DB120".Static_18 OR "DB120".Static_19 OR "DB120".Static_20 OR "DB120".Static_24;
END_REGION

REGION Network 58
   RUNG wire#powerrail
      Contact( "DB120".Static_33 )
      wire#w1
      Coil( #Temp_8 )
   END_RUNG
   RUNG wire#powerrail
      Contact( "DB120".Static_34 )
   END_RUNG wire#w1
   RUNG wire#powerrail
      Contact( "DB120".Static_35 )
   END_RUNG wire#w1
   RUNG wire#powerrail
      Contact( "DB120".Static_36 )
   END_RUNG wire#w1
   RUNG wire#powerrail
      Contact( "DB120".Static_40 )
   END_RUNG wire#w1
   // the same network as SCL:
   #Temp_8 := "DB120".Static_33 OR "DB120".Static_34 OR "DB120".Static_35 OR "DB120".Static_36 OR "DB120".Static_40;
END_REGION

REGION Network 59
   RUNG wire#powerrail
      Contact( "DB120".Static_49 )
      wire#w1
      Coil( #Temp_9 )
   END_RUNG
   RUNG wire#powerrail
      Contact( "DB120".Static_50 )
   END_RUNG wire#w1
   RUNG wire#powerrail
      Contact( "DB120".Static_51 )
   END_RUNG wire#w1
   RUNG wire#powerrail
      Contact( "DB120".Static_52 )
   END_RUNG wire#w1
   RUNG wire#powerrail
      Contact( "DB120".Static_56 )
   END_RUNG wire#w1
   // the same network as SCL:
   #Temp_9 := "DB120".Static_49 OR "DB120".Static_50 OR "DB120".Static_51 OR "DB120".Static_52 OR "DB120".Static_56;
END_REGION

REGION Network 60
